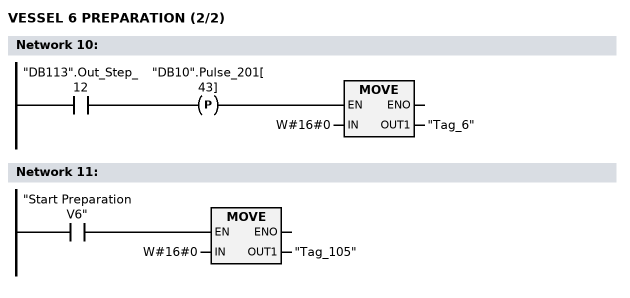
   RUNG wire#powerrail
      Contact( "DB113".Out_Step_12 )
      P_Trig( "DB10".Pulse_201[43] )
      Move(in := W#16#0, out1 => "Tag_6")
   END_RUNG
   // the same network as SCL:
   #_w1 := "DB113".Out_Step_12 AND NOT "DB10".Pulse_201[43];   // rising edge
   "DB10".Pulse_201[43] := "DB113".Out_Step_12;
   IF #_w1 THEN "Tag_6" := W#16#0; END_IF;
END_REGION

REGION Network 11
   RUNG wire#powerrail
      Contact( "Start Preparation V6" )
      Move(in := W#16#0, out1 => "Tag_105")
   END_RUNG
   // the same network as SCL:
   IF "Start Preparation V6" THEN "Tag_105" := W#16#0; END_IF;
END_REGION
END_FUNCTION

FUNCTION "SEQUENCE V7 PREPARATION" : Void   // FC33, LAD
{ S7_Optimized_Access := 'TRUE' }
VERSION : 0.1
   VAR_TEMP   // added for the SCL form of the ladder/FBD networks
      _w1 : Bool;
      _s5time1 : S5Time;
      _w2 : Bool;
      _s5time2 : S5Time;
   END_VAR
BEGIN

REGION Network 1: Start Preparation
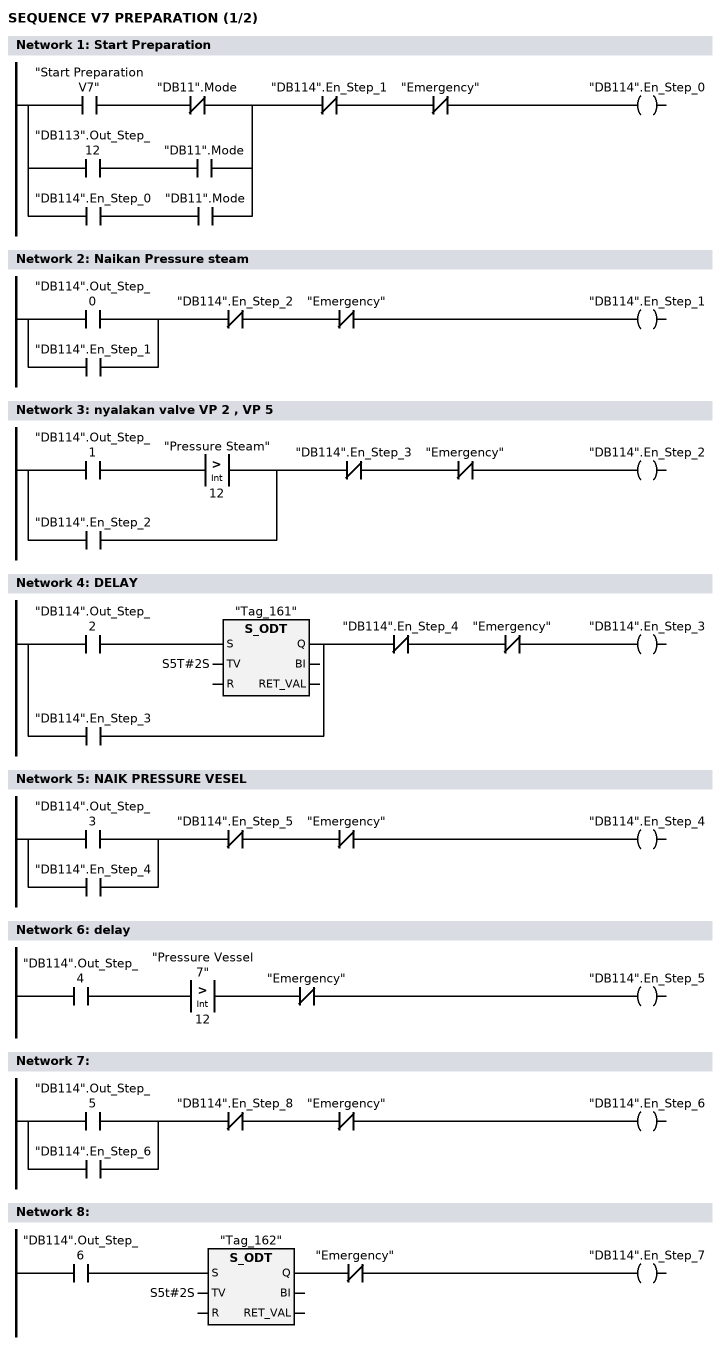
   RUNG wire#powerrail
      Contact( "Start Preparation V7" )
      I_Contact( "DB11".Mode )
      wire#w1
      I_Contact( "DB114".En_Step_1 )
      I_Contact( "Emergency" )
      Coil( "DB114".En_Step_0 )
   END_RUNG
   RUNG wire#powerrail
      Contact( "DB113".Out_Step_12 )
      Contact( "DB11".Mode )
   END_RUNG wire#w1
   RUNG wire#powerrail
      Contact( "DB114".En_Step_0 )
      Contact( "DB11".Mode )
   END_RUNG wire#w1
   // the same network as SCL:
   "DB114".En_Step_0 := (("Start Preparation V7" AND NOT "DB11".Mode) OR ("DB113".Out_Step_12 AND "DB11".Mode) OR ("DB114".En_Step_0 AND "DB11".Mode)) AND NOT "DB114".En_Step_1 AND NOT "Emergency";
END_REGION

REGION Network 2: Naikan Pressure steam
   RUNG wire#powerrail
      Contact( "DB114".Out_Step_0 )
      wire#w1
      I_Contact( "DB114".En_Step_2 )
      I_Contact( "Emergency" )
      Coil( "DB114".En_Step_1 )
   END_RUNG
   RUNG wire#powerrail
      Contact( "DB114".En_Step_1 )
   END_RUNG wire#w1
   // the same network as SCL:
   "DB114".En_Step_1 := ("DB114".Out_Step_0 OR "DB114".En_Step_1) AND NOT "DB114".En_Step_2 AND NOT "Emergency";
END_REGION

REGION Network 3: nyalakan valve VP 2 , VP 5
   RUNG wire#powerrail
      Contact( "DB114".Out_Step_1 )
      { S7_Templates := "SrcType := Int" } GT_Contact(in1 := "Pressure Steam", in2 := 12)
      wire#w1
      I_Contact( "DB114".En_Step_3 )
      I_Contact( "Emergency" )
      Coil( "DB114".En_Step_2 )
   END_RUNG
   RUNG wire#powerrail
      Contact( "DB114".En_Step_2 )
   END_RUNG wire#w1
   // the same network as SCL:
   "DB114".En_Step_2 := (("DB114".Out_Step_1 AND ("Pressure Steam" > 12)) OR "DB114".En_Step_2) AND NOT "DB114".En_Step_3 AND NOT "Emergency";
END_REGION

REGION Network 4: DELAY
   RUNG wire#powerrail
      Contact( "DB114".Out_Step_2 )
      S_ODT(T_NO := "Tag_161", TV := S5T#2S, R :=, BI =>, RET_VAL =>)
      wire#w1
      I_Contact( "DB114".En_Step_4 )
      I_Contact( "Emergency" )
      Coil( "DB114".En_Step_3 )
   END_RUNG
   RUNG wire#powerrail
      Contact( "DB114".En_Step_3 )
   END_RUNG wire#w1
   // the same network as SCL:
   #_s5time1 := S_ODT(T_NO := "Tag_161", S := "DB114".Out_Step_2, TV := S5T#2S, Q => #_w1);
   "DB114".En_Step_3 := (#_w1 OR "DB114".En_Step_3) AND NOT "DB114".En_Step_4 AND NOT "Emergency";
END_REGION

REGION Network 5: NAIK PRESSURE VESEL
   RUNG wire#powerrail
      Contact( "DB114".Out_Step_3 )
      wire#w1
      I_Contact( "DB114".En_Step_5 )
      I_Contact( "Emergency" )
      Coil( "DB114".En_Step_4 )
   END_RUNG
   RUNG wire#powerrail
      Contact( "DB114".En_Step_4 )
   END_RUNG wire#w1
   // the same network as SCL:
   "DB114".En_Step_4 := ("DB114".Out_Step_3 OR "DB114".En_Step_4) AND NOT "DB114".En_Step_5 AND NOT "Emergency";
END_REGION

REGION Network 6: delay
   RUNG wire#powerrail
      Contact( "DB114".Out_Step_4 )
      { S7_Templates := "SrcType := Int" } GT_Contact(in1 := "Pressure Vessel 7", in2 := 12)
      I_Contact( "Emergency" )
      Coil( "DB114".En_Step_5 )
   END_RUNG
   // the same network as SCL:
   "DB114".En_Step_5 := "DB114".Out_Step_4 AND ("Pressure Vessel 7" > 12) AND NOT "Emergency";
END_REGION

REGION Network 7
   RUNG wire#powerrail
      Contact( "DB114".Out_Step_5 )
      wire#w1
      I_Contact( "DB114".En_Step_8 )
      I_Contact( "Emergency" )
      Coil( "DB114".En_Step_6 )
   END_RUNG
   RUNG wire#powerrail
      Contact( "DB114".En_Step_6 )
   END_RUNG wire#w1
   // the same network as SCL:
   "DB114".En_Step_6 := ("DB114".Out_Step_5 OR "DB114".En_Step_6) AND NOT "DB114".En_Step_8 AND NOT "Emergency";
END_REGION

REGION Network 8
   RUNG wire#powerrail
      Contact( "DB114".Out_Step_6 )
      S_ODT(T_NO := "Tag_162", TV := S5t#2S, R :=, BI =>, RET_VAL =>)
      I_Contact( "Emergency" )
      Coil( "DB114".En_Step_7 )
   END_RUNG
   // the same network as SCL:
   #_s5time1 := S_ODT(T_NO := "Tag_162", S := "DB114".Out_Step_6, TV := S5t#2S, Q => #_w1);
   "DB114".En_Step_7 := #_w1 AND NOT "Emergency";
END_REGION

REGION Network 9: TURUNKAN PRESSURE
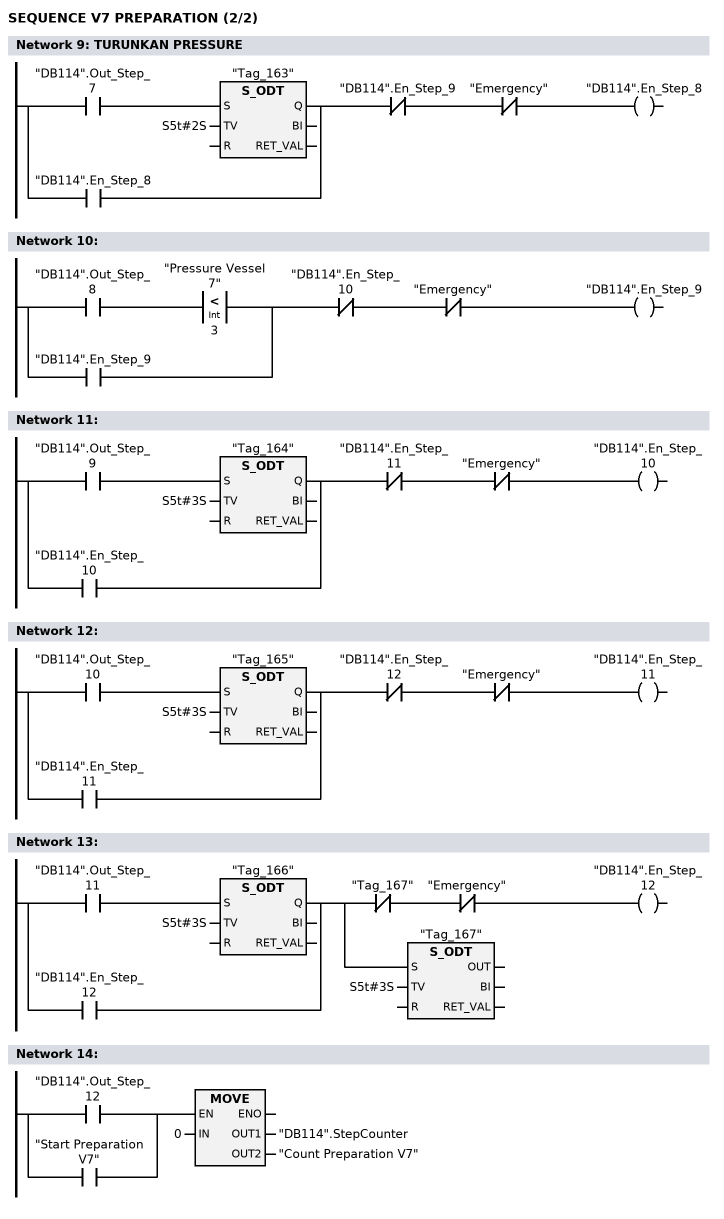
   RUNG wire#powerrail
      Contact( "DB114".Out_Step_7 )
      S_ODT(T_NO := "Tag_163", TV := S5t#2S, R :=, BI =>, RET_VAL =>)
      wire#w1
      I_Contact( "DB114".En_Step_9 )
      I_Contact( "Emergency" )
      Coil( "DB114".En_Step_8 )
   END_RUNG
   RUNG wire#powerrail
      Contact( "DB114".En_Step_8 )
   END_RUNG wire#w1
   // the same network as SCL:
   #_s5time1 := S_ODT(T_NO := "Tag_163", S := "DB114".Out_Step_7, TV := S5t#2S, Q => #_w1);
   "DB114".En_Step_8 := (#_w1 OR "DB114".En_Step_8) AND NOT "DB114".En_Step_9 AND NOT "Emergency";
END_REGION

REGION Network 10
   RUNG wire#powerrail
      Contact( "DB114".Out_Step_8 )
      { S7_Templates := "SrcType := Int" } LT_Contact(in1 := "Pressure Vessel 7", in2 := 3)
      wire#w1
      I_Contact( "DB114".En_Step_10 )
      I_Contact( "Emergency" )
      Coil( "DB114".En_Step_9 )
   END_RUNG
   RUNG wire#powerrail
      Contact( "DB114".En_Step_9 )
   END_RUNG wire#w1
   // the same network as SCL:
   "DB114".En_Step_9 := (("DB114".Out_Step_8 AND ("Pressure Vessel 7" < 3)) OR "DB114".En_Step_9) AND NOT "DB114".En_Step_10 AND NOT "Emergency";
END_REGION

REGION Network 11
   RUNG wire#powerrail
      Contact( "DB114".Out_Step_9 )
      S_ODT(T_NO := "Tag_164", TV := S5t#3S, R :=, BI =>, RET_VAL =>)
      wire#w1
      I_Contact( "DB114".En_Step_11 )
      I_Contact( "Emergency" )
      Coil( "DB114".En_Step_10 )
   END_RUNG
   RUNG wire#powerrail
      Contact( "DB114".En_Step_10 )
   END_RUNG wire#w1
   // the same network as SCL:
   #_s5time1 := S_ODT(T_NO := "Tag_164", S := "DB114".Out_Step_9, TV := S5t#3S, Q => #_w1);
   "DB114".En_Step_10 := (#_w1 OR "DB114".En_Step_10) AND NOT "DB114".En_Step_11 AND NOT "Emergency";
END_REGION

REGION Network 12
   RUNG wire#powerrail
      Contact( "DB114".Out_Step_10 )
      S_ODT(T_NO := "Tag_165", TV := S5t#3S, R :=, BI =>, RET_VAL =>)
      wire#w1
      I_Contact( "DB114".En_Step_12 )
      I_Contact( "Emergency" )
      Coil( "DB114".En_Step_11 )
   END_RUNG
   RUNG wire#powerrail
      Contact( "DB114".En_Step_11 )
   END_RUNG wire#w1
   // the same network as SCL:
   #_s5time1 := S_ODT(T_NO := "Tag_165", S := "DB114".Out_Step_10, TV := S5t#3S, Q => #_w1);
   "DB114".En_Step_11 := (#_w1 OR "DB114".En_Step_11) AND NOT "DB114".En_Step_12 AND NOT "Emergency";
END_REGION

REGION Network 13
   RUNG wire#powerrail
      Contact( "DB114".Out_Step_11 )
      S_ODT(T_NO := "Tag_166", TV := S5t#3S, R :=, BI =>, RET_VAL =>)
      wire#w1
      I_Contact( "Tag_167" )
      I_Contact( "Emergency" )
      Coil( "DB114".En_Step_12 )
   END_RUNG
   RUNG wire#powerrail
      Contact( "DB114".En_Step_12 )
   END_RUNG wire#w1
   RUNG wire#w1
      S_ODT(T_NO := "Tag_167", TV := S5t#3S, R :=, BI =>, RET_VAL =>)
   END_RUNG
   // the same network as SCL:
   #_s5time1 := S_ODT(T_NO := "Tag_166", S := "DB114".Out_Step_11, TV := S5t#3S, Q => #_w1);
   #_w2 := #_w1 OR "DB114".En_Step_12;
   "DB114".En_Step_12 := #_w2 AND NOT "Tag_167" AND NOT "Emergency";
   #_s5time2 := S_ODT(T_NO := "Tag_167", S := #_w2, TV := S5t#3S);
END_REGION

REGION Network 14
   RUNG wire#powerrail
      Contact( "DB114".Out_Step_12 )
      wire#w1
      Move(in := 0, out1 => "DB114".StepCounter, out2 => "Count Preparation V7")
   END_RUNG
   RUNG wire#powerrail
      Contact( "Start Preparation V7" )
   END_RUNG wire#w1
   // the same network as SCL:
   IF "DB114".Out_Step_12 OR "Start Preparation V7" THEN
       "DB114".StepCounter := 0;
       "Count Preparation V7" := 0;
   END_IF;
END_REGION
END_FUNCTION

FUNCTION "VESSEL 7 PREPARATION" : Void   // FC34, LAD
{ S7_Optimized_Access := 'TRUE' }
VERSION : 0.1
   VAR_TEMP   // added for the SCL form of the ladder/FBD networks
      _w1 : Bool;
      _w2 : Bool;
      _w3 : Bool;
      _w4 : Bool;
   END_VAR
BEGIN

REGION Network 1: NAIKAN PRESSURE STEAM
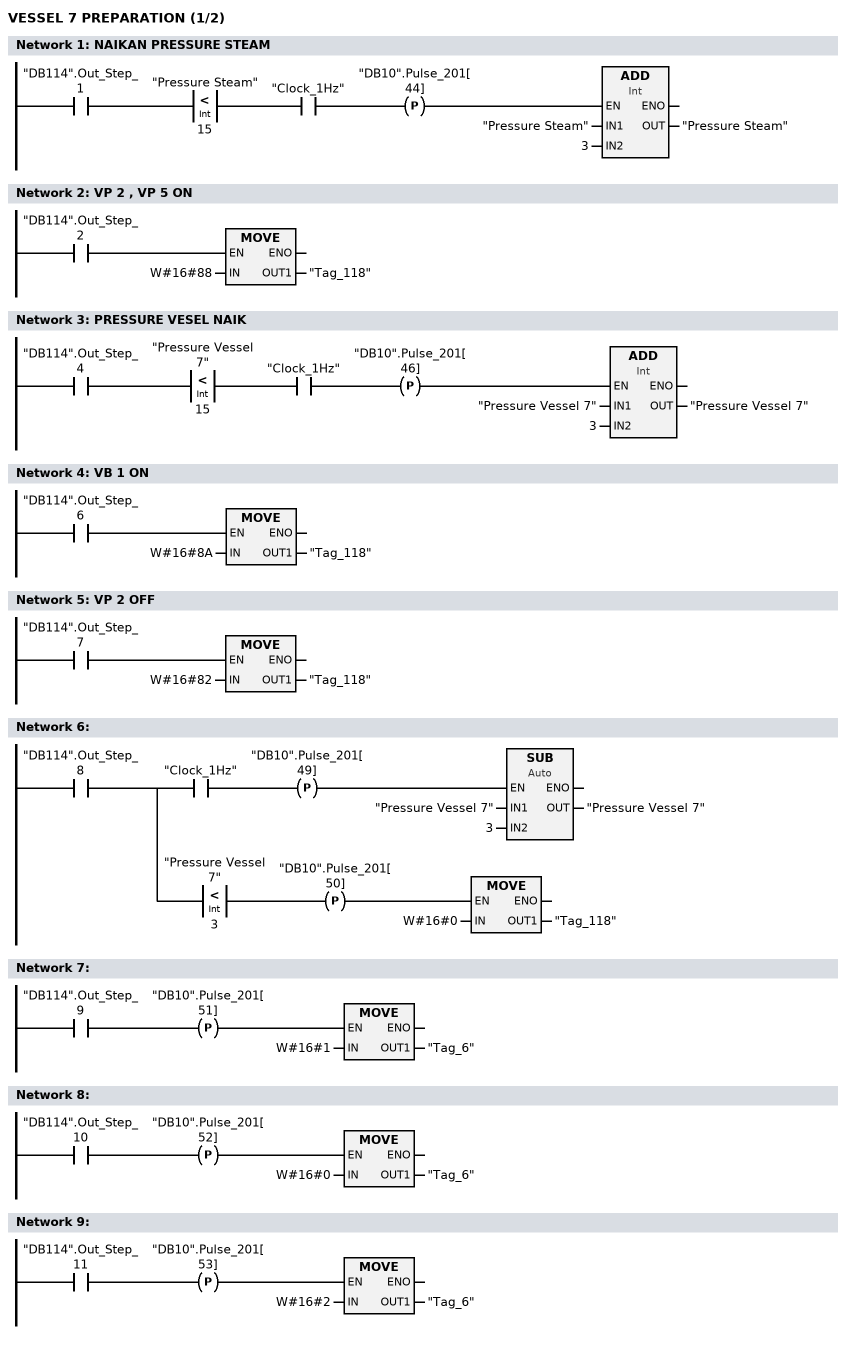
   RUNG wire#powerrail
      Contact( "DB114".Out_Step_1 )
      { S7_Templates := "SrcType := Int" } LT_Contact(in1 := "Pressure Steam", in2 := 15)
      Contact( "Clock_1Hz" )
      P_Trig( "DB10".Pulse_201[44] )
      { S7_Templates := "SrcType := Int" } Add(in1 := "Pressure Steam", in2 := 3, out => "Pressure Steam")
   END_RUNG
   // the same network as SCL:
   #_w1 := "DB114".Out_Step_1 AND ("Pressure Steam" < 15) AND "Clock_1Hz";
   #_w2 := #_w1 AND NOT "DB10".Pulse_201[44];   // rising edge
   "DB10".Pulse_201[44] := #_w1;
   IF #_w2 THEN "Pressure Steam" := "Pressure Steam" + 3; END_IF;
END_REGION

REGION Network 2: VP 2 , VP 5 ON
   RUNG wire#powerrail
      Contact( "DB114".Out_Step_2 )
      Move(in := W#16#88, out1 => "Tag_118")
   END_RUNG
   // the same network as SCL:
   IF "DB114".Out_Step_2 THEN "Tag_118" := W#16#88; END_IF;
END_REGION

REGION Network 3: PRESSURE VESEL NAIK
   RUNG wire#powerrail
      Contact( "DB114".Out_Step_4 )
      { S7_Templates := "SrcType := Int" } LT_Contact(in1 := "Pressure Vessel 7", in2 := 15)
      Contact( "Clock_1Hz" )
      P_Trig( "DB10".Pulse_201[46] )
      { S7_Templates := "SrcType := Int" } Add(in1 := "Pressure Vessel 7", in2 := 3, out => "Pressure Vessel 7")
   END_RUNG
   // the same network as SCL:
   #_w1 := "DB114".Out_Step_4 AND ("Pressure Vessel 7" < 15) AND "Clock_1Hz";
   #_w2 := #_w1 AND NOT "DB10".Pulse_201[46];   // rising edge
   "DB10".Pulse_201[46] := #_w1;
   IF #_w2 THEN "Pressure Vessel 7" := "Pressure Vessel 7" + 3; END_IF;
END_REGION

REGION Network 4: VB 1 ON
   RUNG wire#powerrail
      Contact( "DB114".Out_Step_6 )
      Move(in := W#16#8A, out1 => "Tag_118")
   END_RUNG
   // the same network as SCL:
   IF "DB114".Out_Step_6 THEN "Tag_118" := W#16#8A; END_IF;
END_REGION

REGION Network 5: VP 2 OFF
   RUNG wire#powerrail
      Contact( "DB114".Out_Step_7 )
      Move(in := W#16#82, out1 => "Tag_118")
   END_RUNG
   // the same network as SCL:
   IF "DB114".Out_Step_7 THEN "Tag_118" := W#16#82; END_IF;
END_REGION

REGION Network 6
   RUNG wire#powerrail
      Contact( "DB114".Out_Step_8 )
      wire#w1
      Contact( "Clock_1Hz" )
      P_Trig( "DB10".Pulse_201[49] )
      Sub(in1 := "Pressure Vessel 7", in2 := 3, out => "Pressure Vessel 7")
   END_RUNG
   RUNG wire#w1
      { S7_Templates := "SrcType := Int" } LT_Contact(in1 := "Pressure Vessel 7", in2 := 3)
      P_Trig( "DB10".Pulse_201[50] )
      Move(in := W#16#0, out1 => "Tag_118")
   END_RUNG
   // the same network as SCL:
   #_w1 := "DB114".Out_Step_8 AND "Clock_1Hz";
   #_w2 := #_w1 AND NOT "DB10".Pulse_201[49];   // rising edge
   "DB10".Pulse_201[49] := #_w1;
   IF #_w2 THEN "Pressure Vessel 7" := "Pressure Vessel 7" - 3; END_IF;
   #_w3 := "DB114".Out_Step_8 AND ("Pressure Vessel 7" < 3);
   #_w4 := #_w3 AND NOT "DB10".Pulse_201[50];   // rising edge
   "DB10".Pulse_201[50] := #_w3;
   IF #_w4 THEN "Tag_118" := W#16#0; END_IF;
END_REGION

REGION Network 7
   RUNG wire#powerrail
      Contact( "DB114".Out_Step_9 )
      P_Trig( "DB10".Pulse_201[51] )
      Move(in := W#16#1, out1 => "Tag_6")
   END_RUNG
   // the same network as SCL:
   #_w1 := "DB114".Out_Step_9 AND NOT "DB10".Pulse_201[51];   // rising edge
   "DB10".Pulse_201[51] := "DB114".Out_Step_9;
   IF #_w1 THEN "Tag_6" := W#16#1; END_IF;
END_REGION

REGION Network 8
   RUNG wire#powerrail
      Contact( "DB114".Out_Step_10 )
      P_Trig( "DB10".Pulse_201[52] )
      Move(in := W#16#0, out1 => "Tag_6")
   END_RUNG
   // the same network as SCL:
   #_w1 := "DB114".Out_Step_10 AND NOT "DB10".Pulse_201[52];   // rising edge
   "DB10".Pulse_201[52] := "DB114".Out_Step_10;
   IF #_w1 THEN "Tag_6" := W#16#0; END_IF;
END_REGION

REGION Network 9
   RUNG wire#powerrail
      Contact( "DB114".Out_Step_11 )
      P_Trig( "DB10".Pulse_201[53] )
      Move(in := W#16#2, out1 => "Tag_6")
   END_RUNG
   // the same network as SCL:
   #_w1 := "DB114".Out_Step_11 AND NOT "DB10".Pulse_201[53];   // rising edge
   "DB10".Pulse_201[53] := "DB114".Out_Step_11;
   IF #_w1 THEN "Tag_6" := W#16#2; END_IF;
END_REGION

REGION Network 10
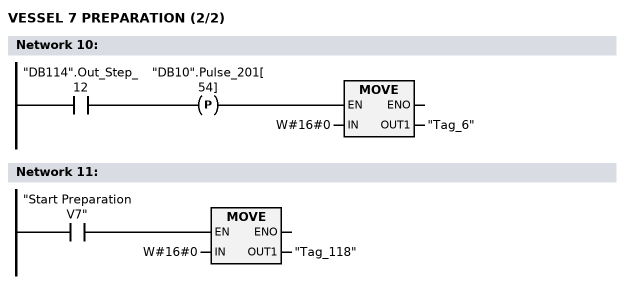
   RUNG wire#powerrail
      Contact( "DB114".Out_Step_12 )
      P_Trig( "DB10".Pulse_201[54] )
      Move(in := W#16#0, out1 => "Tag_6")
   END_RUNG
   // the same network as SCL:
   #_w1 := "DB114".Out_Step_12 AND NOT "DB10".Pulse_201[54];   // rising edge
   "DB10".Pulse_201[54] := "DB114".Out_Step_12;
   IF #_w1 THEN "Tag_6" := W#16#0; END_IF;
END_REGION

REGION Network 11
   RUNG wire#powerrail
      Contact( "Start Preparation V7" )
      Move(in := W#16#0, out1 => "Tag_118")
   END_RUNG
   // the same network as SCL:
   IF "Start Preparation V7" THEN "Tag_118" := W#16#0; END_IF;
END_REGION
END_FUNCTION

FUNCTION "SEQUENCE CLEAN" : Void   // FC35, LAD
{ S7_Optimized_Access := 'TRUE' }
VERSION : 0.1
   VAR_TEMP   // added for the SCL form of the ladder/FBD networks
      _w1 : Bool;
      _w2 : Bool;
      _s5time1 : S5Time;
   END_VAR
BEGIN

REGION Network 1
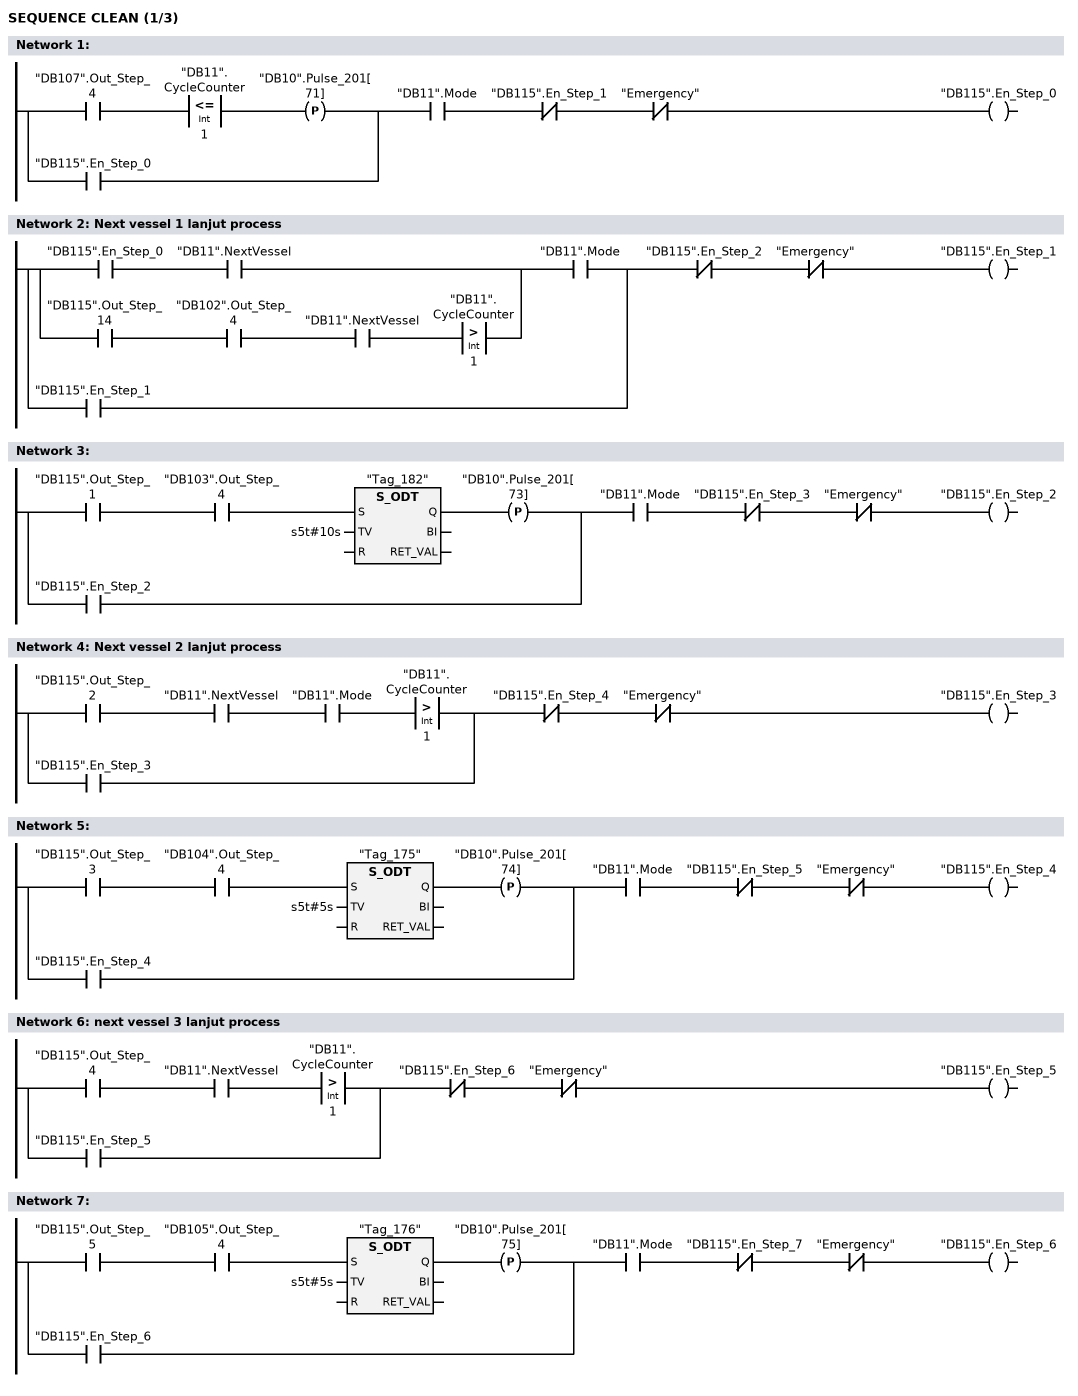
   RUNG wire#powerrail
      Contact( "DB107".Out_Step_4 )
      { S7_Templates := "SrcType := Int" } LE_Contact(in1 := "DB11".CycleCounter, in2 := 1)
      P_Trig( "DB10".Pulse_201[71] )
      wire#w1
      Contact( "DB11".Mode )
      I_Contact( "DB115".En_Step_1 )
      I_Contact( "Emergency" )
      Coil( "DB115".En_Step_0 )
   END_RUNG
   RUNG wire#powerrail
      Contact( "DB115".En_Step_0 )
   END_RUNG wire#w1
   // the same network as SCL:
   #_w1 := "DB107".Out_Step_4 AND ("DB11".CycleCounter <= 1);
   #_w2 := #_w1 AND NOT "DB10".Pulse_201[71];   // rising edge
   "DB10".Pulse_201[71] := #_w1;
   "DB115".En_Step_0 := (#_w2 OR "DB115".En_Step_0) AND "DB11".Mode AND NOT "DB115".En_Step_1 AND NOT "Emergency";
END_REGION

REGION Network 2: Next vessel 1 lanjut process
   RUNG wire#powerrail
      Contact( "DB115".En_Step_0 )
      Contact( "DB11".NextVessel )
      wire#w1
      Contact( "DB11".Mode )
      wire#w2
      I_Contact( "DB115".En_Step_2 )
      I_Contact( "Emergency" )
      Coil( "DB115".En_Step_1 )
   END_RUNG
   RUNG wire#powerrail
      Contact( "DB115".Out_Step_14 )
      Contact( "DB102".Out_Step_4 )
      Contact( "DB11".NextVessel )
      { S7_Templates := "SrcType := Int" } GT_Contact(in1 := "DB11".CycleCounter, in2 := 1)
   END_RUNG wire#w1
   RUNG wire#powerrail
      Contact( "DB115".En_Step_1 )
   END_RUNG wire#w2
   // the same network as SCL:
   "DB115".En_Step_1 := (((("DB115".En_Step_0 AND "DB11".NextVessel) OR ("DB115".Out_Step_14 AND "DB102".Out_Step_4 AND "DB11".NextVessel AND ("DB11".CycleCounter > 1))) AND "DB11".Mode) OR "DB115".En_Step_1) AND NOT "DB115".En_Step_2 AND NOT "Emergency";
END_REGION

REGION Network 3
   RUNG wire#powerrail
      Contact( "DB115".Out_Step_1 )
      Contact( "DB103".Out_Step_4 )
      S_ODT(T_NO := "Tag_182", TV := s5t#10s, R :=, BI =>, RET_VAL =>)
      P_Trig( "DB10".Pulse_201[73] )
      wire#w1
      Contact( "DB11".Mode )
      I_Contact( "DB115".En_Step_3 )
      I_Contact( "Emergency" )
      Coil( "DB115".En_Step_2 )
   END_RUNG
   RUNG wire#powerrail
      Contact( "DB115".En_Step_2 )
   END_RUNG wire#w1
   // the same network as SCL:
   #_s5time1 := S_ODT(T_NO := "Tag_182",
                      S := "DB115".Out_Step_1 AND "DB103".Out_Step_4,
                      TV := s5t#10s,
                      Q => #_w1);
   #_w2 := #_w1 AND NOT "DB10".Pulse_201[73];   // rising edge
   "DB10".Pulse_201[73] := #_w1;
   "DB115".En_Step_2 := (#_w2 OR "DB115".En_Step_2) AND "DB11".Mode AND NOT "DB115".En_Step_3 AND NOT "Emergency";
END_REGION

REGION Network 4: Next vessel 2 lanjut process
   RUNG wire#powerrail
      Contact( "DB115".Out_Step_2 )
      Contact( "DB11".NextVessel )
      Contact( "DB11".Mode )
      { S7_Templates := "SrcType := Int" } GT_Contact(in1 := "DB11".CycleCounter, in2 := 1)
      wire#w1
      I_Contact( "DB115".En_Step_4 )
      I_Contact( "Emergency" )
      Coil( "DB115".En_Step_3 )
   END_RUNG
   RUNG wire#powerrail
      Contact( "DB115".En_Step_3 )
   END_RUNG wire#w1
   // the same network as SCL:
   "DB115".En_Step_3 := (("DB115".Out_Step_2 AND "DB11".NextVessel AND "DB11".Mode AND ("DB11".CycleCounter > 1)) OR "DB115".En_Step_3) AND NOT "DB115".En_Step_4 AND NOT "Emergency";
END_REGION

REGION Network 5
   RUNG wire#powerrail
      Contact( "DB115".Out_Step_3 )
      Contact( "DB104".Out_Step_4 )
      S_ODT(T_NO := "Tag_175", TV := s5t#5s, R :=, BI =>, RET_VAL =>)
      P_Trig( "DB10".Pulse_201[74] )
      wire#w1
      Contact( "DB11".Mode )
      I_Contact( "DB115".En_Step_5 )
      I_Contact( "Emergency" )
      Coil( "DB115".En_Step_4 )
   END_RUNG
   RUNG wire#powerrail
      Contact( "DB115".En_Step_4 )
   END_RUNG wire#w1
   // the same network as SCL:
   #_s5time1 := S_ODT(T_NO := "Tag_175",
                      S := "DB115".Out_Step_3 AND "DB104".Out_Step_4,
                      TV := s5t#5s,
                      Q => #_w1);
   #_w2 := #_w1 AND NOT "DB10".Pulse_201[74];   // rising edge
   "DB10".Pulse_201[74] := #_w1;
   "DB115".En_Step_4 := (#_w2 OR "DB115".En_Step_4) AND "DB11".Mode AND NOT "DB115".En_Step_5 AND NOT "Emergency";
END_REGION

REGION Network 6: next vessel 3 lanjut process
   RUNG wire#powerrail
      Contact( "DB115".Out_Step_4 )
      Contact( "DB11".NextVessel )
      { S7_Templates := "SrcType := Int" } GT_Contact(in1 := "DB11".CycleCounter, in2 := 1)
      wire#w1
      I_Contact( "DB115".En_Step_6 )
      I_Contact( "Emergency" )
      Coil( "DB115".En_Step_5 )
   END_RUNG
   RUNG wire#powerrail
      Contact( "DB115".En_Step_5 )
   END_RUNG wire#w1
   // the same network as SCL:
   "DB115".En_Step_5 := (("DB115".Out_Step_4 AND "DB11".NextVessel AND ("DB11".CycleCounter > 1)) OR "DB115".En_Step_5) AND NOT "DB115".En_Step_6 AND NOT "Emergency";
END_REGION

REGION Network 7
   RUNG wire#powerrail
      Contact( "DB115".Out_Step_5 )
      Contact( "DB105".Out_Step_4 )
      S_ODT(T_NO := "Tag_176", TV := s5t#5s, R :=, BI =>, RET_VAL =>)
      P_Trig( "DB10".Pulse_201[75] )
      wire#w1
      Contact( "DB11".Mode )
      I_Contact( "DB115".En_Step_7 )
      I_Contact( "Emergency" )
      Coil( "DB115".En_Step_6 )
   END_RUNG
   RUNG wire#powerrail
      Contact( "DB115".En_Step_6 )
   END_RUNG wire#w1
   // the same network as SCL:
   #_s5time1 := S_ODT(T_NO := "Tag_176",
                      S := "DB115".Out_Step_5 AND "DB105".Out_Step_4,
                      TV := s5t#5s,
                      Q => #_w1);
   #_w2 := #_w1 AND NOT "DB10".Pulse_201[75];   // rising edge
   "DB10".Pulse_201[75] := #_w1;
   "DB115".En_Step_6 := (#_w2 OR "DB115".En_Step_6) AND "DB11".Mode AND NOT "DB115".En_Step_7 AND NOT "Emergency";
END_REGION

REGION Network 8: next vessel 4 lanjut process
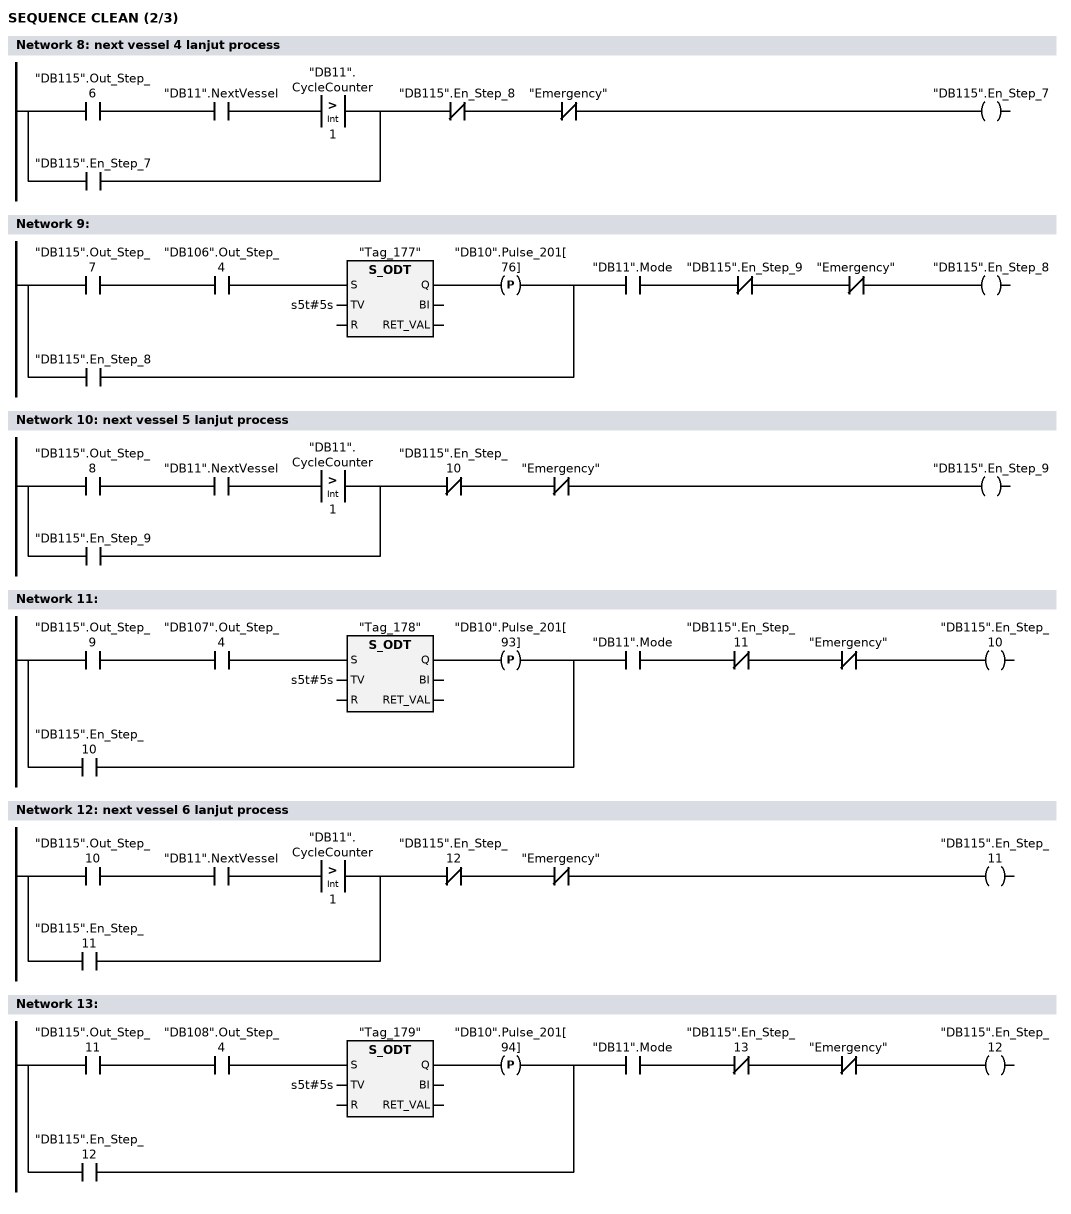
   RUNG wire#powerrail
      Contact( "DB115".Out_Step_6 )
      Contact( "DB11".NextVessel )
      { S7_Templates := "SrcType := Int" } GT_Contact(in1 := "DB11".CycleCounter, in2 := 1)
      wire#w1
      I_Contact( "DB115".En_Step_8 )
      I_Contact( "Emergency" )
      Coil( "DB115".En_Step_7 )
   END_RUNG
   RUNG wire#powerrail
      Contact( "DB115".En_Step_7 )
   END_RUNG wire#w1
   // the same network as SCL:
   "DB115".En_Step_7 := (("DB115".Out_Step_6 AND "DB11".NextVessel AND ("DB11".CycleCounter > 1)) OR "DB115".En_Step_7) AND NOT "DB115".En_Step_8 AND NOT "Emergency";
END_REGION

REGION Network 9
   RUNG wire#powerrail
      Contact( "DB115".Out_Step_7 )
      Contact( "DB106".Out_Step_4 )
      S_ODT(T_NO := "Tag_177", TV := s5t#5s, R :=, BI =>, RET_VAL =>)
      P_Trig( "DB10".Pulse_201[76] )
      wire#w1
      Contact( "DB11".Mode )
      I_Contact( "DB115".En_Step_9 )
      I_Contact( "Emergency" )
      Coil( "DB115".En_Step_8 )
   END_RUNG
   RUNG wire#powerrail
      Contact( "DB115".En_Step_8 )
   END_RUNG wire#w1
   // the same network as SCL:
   #_s5time1 := S_ODT(T_NO := "Tag_177",
                      S := "DB115".Out_Step_7 AND "DB106".Out_Step_4,
                      TV := s5t#5s,
                      Q => #_w1);
   #_w2 := #_w1 AND NOT "DB10".Pulse_201[76];   // rising edge
   "DB10".Pulse_201[76] := #_w1;
   "DB115".En_Step_8 := (#_w2 OR "DB115".En_Step_8) AND "DB11".Mode AND NOT "DB115".En_Step_9 AND NOT "Emergency";
END_REGION

REGION Network 10: next vessel 5 lanjut process
   RUNG wire#powerrail
      Contact( "DB115".Out_Step_8 )
      Contact( "DB11".NextVessel )
      { S7_Templates := "SrcType := Int" } GT_Contact(in1 := "DB11".CycleCounter, in2 := 1)
      wire#w1
      I_Contact( "DB115".En_Step_10 )
      I_Contact( "Emergency" )
      Coil( "DB115".En_Step_9 )
   END_RUNG
   RUNG wire#powerrail
      Contact( "DB115".En_Step_9 )
   END_RUNG wire#w1
   // the same network as SCL:
   "DB115".En_Step_9 := (("DB115".Out_Step_8 AND "DB11".NextVessel AND ("DB11".CycleCounter > 1)) OR "DB115".En_Step_9) AND NOT "DB115".En_Step_10 AND NOT "Emergency";
END_REGION

REGION Network 11
   RUNG wire#powerrail
      Contact( "DB115".Out_Step_9 )
      Contact( "DB107".Out_Step_4 )
      S_ODT(T_NO := "Tag_178", TV := s5t#5s, R :=, BI =>, RET_VAL =>)
      P_Trig( "DB10".Pulse_201[93] )
      wire#w1
      Contact( "DB11".Mode )
      I_Contact( "DB115".En_Step_11 )
      I_Contact( "Emergency" )
      Coil( "DB115".En_Step_10 )
   END_RUNG
   RUNG wire#powerrail
      Contact( "DB115".En_Step_10 )
   END_RUNG wire#w1
   // the same network as SCL:
   #_s5time1 := S_ODT(T_NO := "Tag_178",
                      S := "DB115".Out_Step_9 AND "DB107".Out_Step_4,
                      TV := s5t#5s,
                      Q => #_w1);
   #_w2 := #_w1 AND NOT "DB10".Pulse_201[93];   // rising edge
   "DB10".Pulse_201[93] := #_w1;
   "DB115".En_Step_10 := (#_w2 OR "DB115".En_Step_10) AND "DB11".Mode AND NOT "DB115".En_Step_11 AND NOT "Emergency";
END_REGION

REGION Network 12: next vessel 6 lanjut process
   RUNG wire#powerrail
      Contact( "DB115".Out_Step_10 )
      Contact( "DB11".NextVessel )
      { S7_Templates := "SrcType := Int" } GT_Contact(in1 := "DB11".CycleCounter, in2 := 1)
      wire#w1
      I_Contact( "DB115".En_Step_12 )
      I_Contact( "Emergency" )
      Coil( "DB115".En_Step_11 )
   END_RUNG
   RUNG wire#powerrail
      Contact( "DB115".En_Step_11 )
   END_RUNG wire#w1
   // the same network as SCL:
   "DB115".En_Step_11 := (("DB115".Out_Step_10 AND "DB11".NextVessel AND ("DB11".CycleCounter > 1)) OR "DB115".En_Step_11) AND NOT "DB115".En_Step_12 AND NOT "Emergency";
END_REGION

REGION Network 13
   RUNG wire#powerrail
      Contact( "DB115".Out_Step_11 )
      Contact( "DB108".Out_Step_4 )
      S_ODT(T_NO := "Tag_179", TV := s5t#5s, R :=, BI =>, RET_VAL =>)
      P_Trig( "DB10".Pulse_201[94] )
      wire#w1
      Contact( "DB11".Mode )
      I_Contact( "DB115".En_Step_13 )
      I_Contact( "Emergency" )
      Coil( "DB115".En_Step_12 )
   END_RUNG
   RUNG wire#powerrail
      Contact( "DB115".En_Step_12 )
   END_RUNG wire#w1
   // the same network as SCL:
   #_s5time1 := S_ODT(T_NO := "Tag_179",
                      S := "DB115".Out_Step_11 AND "DB108".Out_Step_4,
                      TV := s5t#5s,
                      Q => #_w1);
   #_w2 := #_w1 AND NOT "DB10".Pulse_201[94];   // rising edge
   "DB10".Pulse_201[94] := #_w1;
   "DB115".En_Step_12 := (#_w2 OR "DB115".En_Step_12) AND "DB11".Mode AND NOT "DB115".En_Step_13 AND NOT "Emergency";
END_REGION

REGION Network 14: next vessel 7 lanjut process